REGION Network 181
   RUNG wire#powerrail
      Move(in := "Carrier_38_CarrierDriveAlarm", out1 => "DB_SDC_EMS_TA".EMS[38].TA[1].ALARM)
      wire#w1
      Move(in := "Carrier_38_CarrierDriveAlarm", out1 => "EMS".Carrier[38].SDC_IN.CarrierDriveAlarms)
   END_RUNG
   RUNG wire#powerrail
      Contact( "IndiconTempDebugON" )
   END_RUNG wire#w1
   // the same network as SCL:
   "DB_SDC_EMS_TA".EMS[38].TA[1].ALARM := "Carrier_38_CarrierDriveAlarm";
   IF TRUE OR "IndiconTempDebugON" THEN
       "EMS".Carrier[38].SDC_IN.CarrierDriveAlarms := "Carrier_38_CarrierDriveAlarm";
   END_IF;
END_REGION

REGION Network 182
   RUNG wire#powerrail
      Move(in := "Carrier_38_SDCFaultCode", out1 => "DB101_DB_SDC_FAULTS".Carrier_Fault[38])
      wire#w1
      Move(in := "Carrier_38_SDCFaultCode", out1 => "EMS".Carrier[38].SDC_IN.CarrierFaults)
   END_RUNG
   RUNG wire#powerrail
      Contact( "IndiconTempDebugON" )
   END_RUNG wire#w1
   // the same network as SCL:
   "DB101_DB_SDC_FAULTS".Carrier_Fault[38] := "Carrier_38_SDCFaultCode";
   IF TRUE OR "IndiconTempDebugON" THEN
       "EMS".Carrier[38].SDC_IN.CarrierFaults := "Carrier_38_SDCFaultCode";
   END_IF;
END_REGION

REGION Network 183
   RUNG wire#powerrail
      Contact( "Carrier_38_Status.5" )
      Coil( "EMS".Carrier[38].SDC_IN.RunningFWD )
   END_RUNG
   // the same network as SCL:
   "EMS".Carrier[38].SDC_IN.RunningFWD := "Carrier_38_Status.5";
END_REGION

REGION Network 184
   RUNG wire#powerrail
      Contact( "Carrier_38_Status.6" )
      Coil( "EMS".Carrier[38].SDC_IN.RunningREV )
   END_RUNG
   // the same network as SCL:
   "EMS".Carrier[38].SDC_IN.RunningREV := "Carrier_38_Status.6";
END_REGION

REGION Network 185
   RUNG wire#powerrail
      Contact( "Carrier_38_Status.7" )
      Coil( "EMS".Carrier[38].SDC_IN.IR_Remote_9_Pressed )
   END_RUNG
   // the same network as SCL:
   "EMS".Carrier[38].SDC_IN.IR_Remote_9_Pressed := "Carrier_38_Status.7";
END_REGION

REGION Network 186
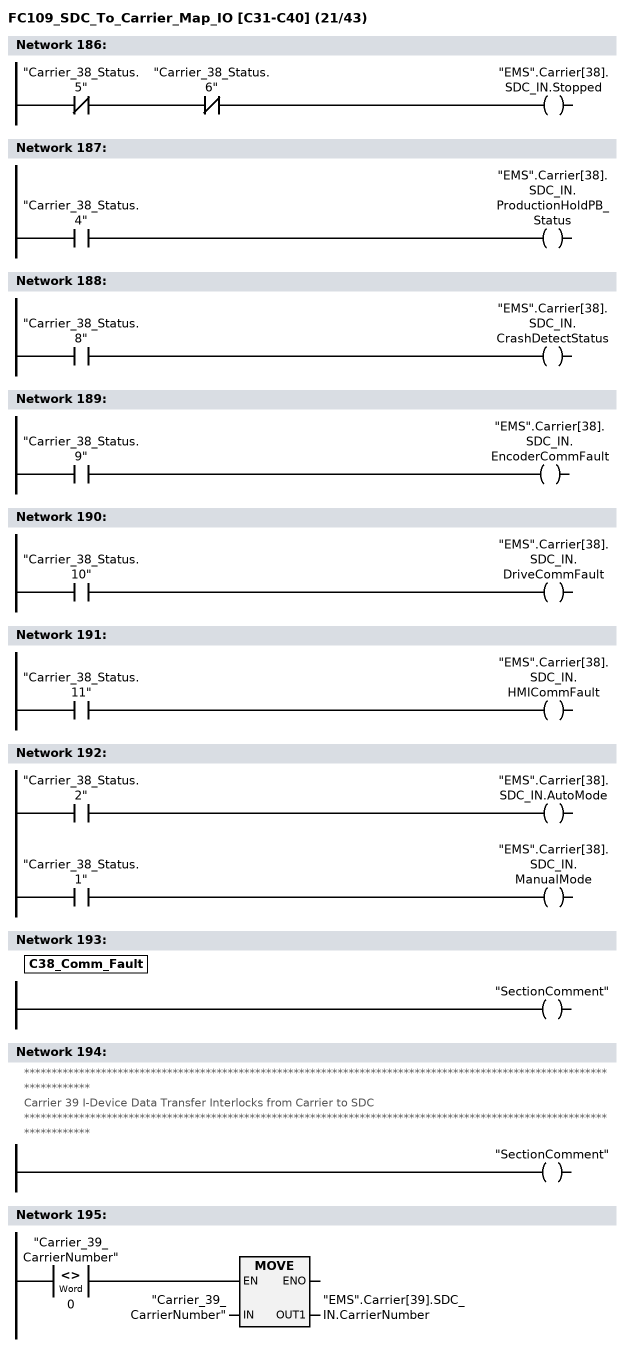
   RUNG wire#powerrail
      I_Contact( "Carrier_38_Status.5" )
      I_Contact( "Carrier_38_Status.6" )
      Coil( "EMS".Carrier[38].SDC_IN.Stopped )
   END_RUNG
   // the same network as SCL:
   "EMS".Carrier[38].SDC_IN.Stopped := NOT "Carrier_38_Status.5" AND NOT "Carrier_38_Status.6";
END_REGION

REGION Network 187
   RUNG wire#powerrail
      Contact( "Carrier_38_Status.4" )
      Coil( "EMS".Carrier[38].SDC_IN.ProductionHoldPB_Status )
   END_RUNG
   // the same network as SCL:
   "EMS".Carrier[38].SDC_IN.ProductionHoldPB_Status := "Carrier_38_Status.4";
END_REGION

REGION Network 188
   RUNG wire#powerrail
      Contact( "Carrier_38_Status.8" )
      Coil( "EMS".Carrier[38].SDC_IN.CrashDetectStatus )
   END_RUNG
   // the same network as SCL:
   "EMS".Carrier[38].SDC_IN.CrashDetectStatus := "Carrier_38_Status.8";
END_REGION

REGION Network 189
   RUNG wire#powerrail
      Contact( "Carrier_38_Status.9" )
      Coil( "EMS".Carrier[38].SDC_IN.EncoderCommFault )
   END_RUNG
   // the same network as SCL:
   "EMS".Carrier[38].SDC_IN.EncoderCommFault := "Carrier_38_Status.9";
END_REGION

REGION Network 190
   RUNG wire#powerrail
      Contact( "Carrier_38_Status.10" )
      Coil( "EMS".Carrier[38].SDC_IN.DriveCommFault )
   END_RUNG
   // the same network as SCL:
   "EMS".Carrier[38].SDC_IN.DriveCommFault := "Carrier_38_Status.10";
END_REGION

REGION Network 191
   RUNG wire#powerrail
      Contact( "Carrier_38_Status.11" )
      Coil( "EMS".Carrier[38].SDC_IN.HMICommFault )
   END_RUNG
   // the same network as SCL:
   "EMS".Carrier[38].SDC_IN.HMICommFault := "Carrier_38_Status.11";
END_REGION

REGION Network 192
   RUNG wire#powerrail
      Contact( "Carrier_38_Status.2" )
      Coil( "EMS".Carrier[38].SDC_IN.AutoMode )
   END_RUNG
   RUNG wire#powerrail
      Contact( "Carrier_38_Status.1" )
      Coil( "EMS".Carrier[38].SDC_IN.ManualMode )
   END_RUNG
   // the same network as SCL:
   "EMS".Carrier[38].SDC_IN.AutoMode := "Carrier_38_Status.2";
   "EMS".Carrier[38].SDC_IN.ManualMode := "Carrier_38_Status.1";
END_REGION

REGION Network 193
   Label( C38_Comm_Fault )
   RUNG wire#powerrail
      Coil( "SectionComment" )
   END_RUNG
   // the same network as SCL:
   C38_Comm_Fault:
   "SectionComment" := TRUE;
END_REGION

REGION Network 194
   // **********************************************************************************************************************
   // 
   // Carrier 39 I-Device Data Transfer Interlocks from Carrier to SDC
   // 
   // **********************************************************************************************************************
   RUNG wire#powerrail
      Coil( "SectionComment" )
   END_RUNG
   // the same network as SCL:
   "SectionComment" := TRUE;
END_REGION

REGION Network 195
   RUNG wire#powerrail
      { S7_Templates := "SrcType := Word" } NE_Contact(in1 := "Carrier_39_CarrierNumber", in2 := 0)
      Move(in := "Carrier_39_CarrierNumber", out1 => "EMS".Carrier[39].SDC_IN.CarrierNumber)
   END_RUNG
   // the same network as SCL:
   IF "Carrier_39_CarrierNumber" <> 0 THEN
       "EMS".Carrier[39].SDC_IN.CarrierNumber := "Carrier_39_CarrierNumber";
   END_IF;
END_REGION

REGION Network 196
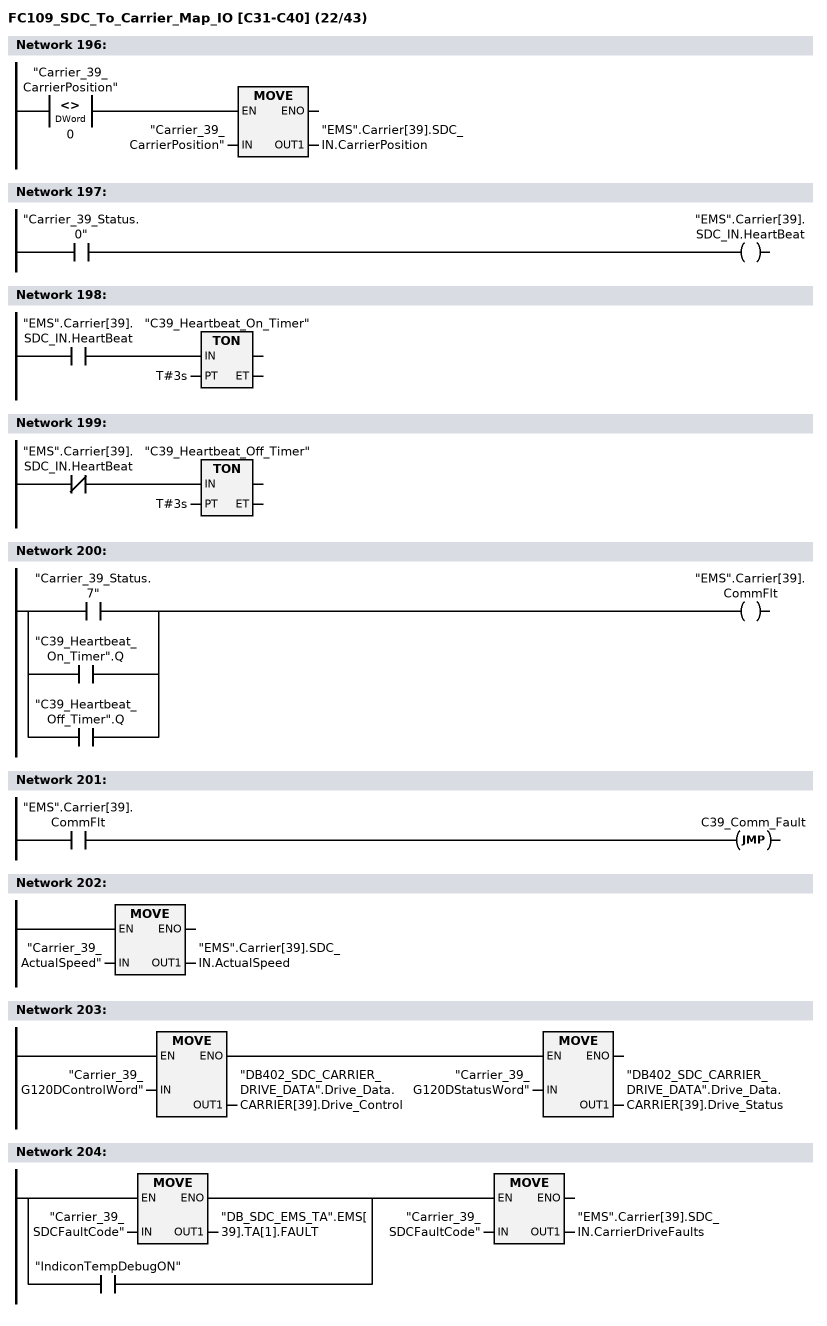
   RUNG wire#powerrail
      { S7_Templates := "SrcType := DWord" } NE_Contact(in1 := "Carrier_39_CarrierPosition", in2 := 0)
      Move(in := "Carrier_39_CarrierPosition", out1 => "EMS".Carrier[39].SDC_IN.CarrierPosition)
   END_RUNG
   // the same network as SCL:
   IF "Carrier_39_CarrierPosition" <> 0 THEN
       "EMS".Carrier[39].SDC_IN.CarrierPosition := "Carrier_39_CarrierPosition";
   END_IF;
END_REGION

REGION Network 197
   RUNG wire#powerrail
      Contact( "Carrier_39_Status.0" )
      Coil( "EMS".Carrier[39].SDC_IN.HeartBeat )
   END_RUNG
   // the same network as SCL:
   "EMS".Carrier[39].SDC_IN.HeartBeat := "Carrier_39_Status.0";
END_REGION

REGION Network 198
   "C39_Heartbeat_On_Timer".TON(IN := "EMS".Carrier[39].SDC_IN.HeartBeat, PT := T#3s);
END_REGION

REGION Network 199
   "C39_Heartbeat_Off_Timer".TON(IN := NOT "EMS".Carrier[39].SDC_IN.HeartBeat, PT := T#3s);
END_REGION

REGION Network 200
   RUNG wire#powerrail
      Contact( "Carrier_39_Status.7" )
      wire#w1
      Coil( "EMS".Carrier[39].CommFlt )
   END_RUNG
   RUNG wire#powerrail
      Contact( "C39_Heartbeat_On_Timer".Q )
   END_RUNG wire#w1
   RUNG wire#powerrail
      Contact( "C39_Heartbeat_Off_Timer".Q )
   END_RUNG wire#w1
   // the same network as SCL:
   "EMS".Carrier[39].CommFlt := "Carrier_39_Status.7" OR "C39_Heartbeat_On_Timer".Q OR "C39_Heartbeat_Off_Timer".Q;
END_REGION

REGION Network 201
   RUNG wire#powerrail
      Contact( "EMS".Carrier[39].CommFlt )
      JumpCoil( C39_Comm_Fault )
   END_RUNG
   // the same network as SCL:
   IF "EMS".Carrier[39].CommFlt THEN GOTO C39_Comm_Fault; END_IF;
END_REGION

REGION Network 202
   RUNG wire#powerrail
      Move(in := "Carrier_39_ActualSpeed", out1 => "EMS".Carrier[39].SDC_IN.ActualSpeed)
   END_RUNG
   // the same network as SCL:
   "EMS".Carrier[39].SDC_IN.ActualSpeed := "Carrier_39_ActualSpeed";
END_REGION

REGION Network 203
   RUNG wire#powerrail
      Move(in := "Carrier_39_G120DControlWord", out1 => "DB402_SDC_CARRIER_DRIVE_DATA".Drive_Data.CARRIER[39].Drive_Control)
      Move(in := "Carrier_39_G120DStatusWord", out1 => "DB402_SDC_CARRIER_DRIVE_DATA".Drive_Data.CARRIER[39].Drive_Status)
   END_RUNG
   // the same network as SCL:
   "DB402_SDC_CARRIER_DRIVE_DATA".Drive_Data.CARRIER[39].Drive_Control := "Carrier_39_G120DControlWord";
   "DB402_SDC_CARRIER_DRIVE_DATA".Drive_Data.CARRIER[39].Drive_Status := "Carrier_39_G120DStatusWord";
END_REGION

REGION Network 204
   RUNG wire#powerrail
      Move(in := "Carrier_39_SDCFaultCode", out1 => "DB_SDC_EMS_TA".EMS[39].TA[1].FAULT)
      wire#w1
      Move(in := "Carrier_39_SDCFaultCode", out1 => "EMS".Carrier[39].SDC_IN.CarrierDriveFaults)
   END_RUNG
   RUNG wire#powerrail
      Contact( "IndiconTempDebugON" )
   END_RUNG wire#w1
   // the same network as SCL:
   "DB_SDC_EMS_TA".EMS[39].TA[1].FAULT := "Carrier_39_SDCFaultCode";
   IF TRUE OR "IndiconTempDebugON" THEN
       "EMS".Carrier[39].SDC_IN.CarrierDriveFaults := "Carrier_39_SDCFaultCode";
   END_IF;
END_REGION

REGION Network 205
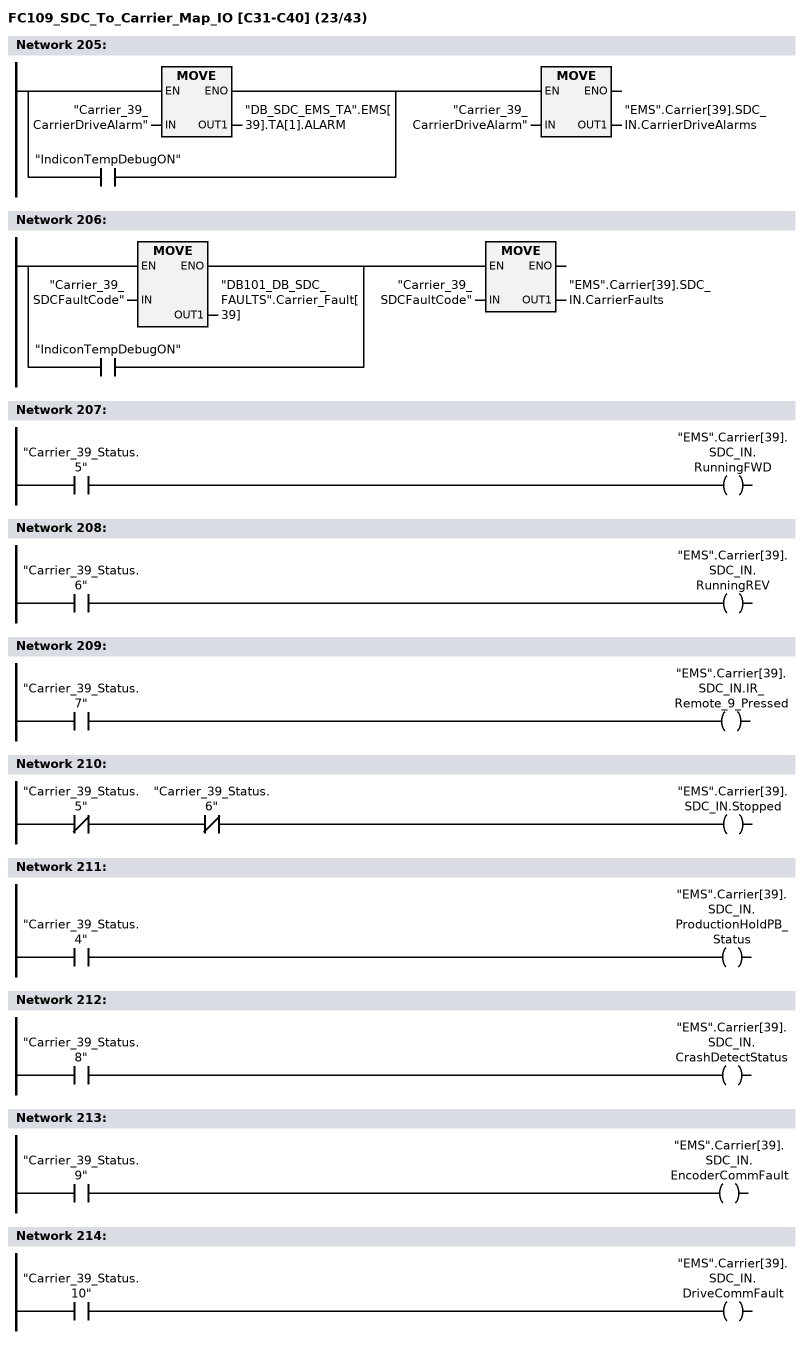
   RUNG wire#powerrail
      Move(in := "Carrier_39_CarrierDriveAlarm", out1 => "DB_SDC_EMS_TA".EMS[39].TA[1].ALARM)
      wire#w1
      Move(in := "Carrier_39_CarrierDriveAlarm", out1 => "EMS".Carrier[39].SDC_IN.CarrierDriveAlarms)
   END_RUNG
   RUNG wire#powerrail
      Contact( "IndiconTempDebugON" )
   END_RUNG wire#w1
   // the same network as SCL:
   "DB_SDC_EMS_TA".EMS[39].TA[1].ALARM := "Carrier_39_CarrierDriveAlarm";
   IF TRUE OR "IndiconTempDebugON" THEN
       "EMS".Carrier[39].SDC_IN.CarrierDriveAlarms := "Carrier_39_CarrierDriveAlarm";
   END_IF;
END_REGION

REGION Network 206
   RUNG wire#powerrail
      Move(in := "Carrier_39_SDCFaultCode", out1 => "DB101_DB_SDC_FAULTS".Carrier_Fault[39])
      wire#w1
      Move(in := "Carrier_39_SDCFaultCode", out1 => "EMS".Carrier[39].SDC_IN.CarrierFaults)
   END_RUNG
   RUNG wire#powerrail
      Contact( "IndiconTempDebugON" )
   END_RUNG wire#w1
   // the same network as SCL:
   "DB101_DB_SDC_FAULTS".Carrier_Fault[39] := "Carrier_39_SDCFaultCode";
   IF TRUE OR "IndiconTempDebugON" THEN
       "EMS".Carrier[39].SDC_IN.CarrierFaults := "Carrier_39_SDCFaultCode";
   END_IF;
END_REGION

REGION Network 207
   RUNG wire#powerrail
      Contact( "Carrier_39_Status.5" )
      Coil( "EMS".Carrier[39].SDC_IN.RunningFWD )
   END_RUNG
   // the same network as SCL:
   "EMS".Carrier[39].SDC_IN.RunningFWD := "Carrier_39_Status.5";
END_REGION

REGION Network 208
   RUNG wire#powerrail
      Contact( "Carrier_39_Status.6" )
      Coil( "EMS".Carrier[39].SDC_IN.RunningREV )
   END_RUNG
   // the same network as SCL:
   "EMS".Carrier[39].SDC_IN.RunningREV := "Carrier_39_Status.6";
END_REGION

REGION Network 209
   RUNG wire#powerrail
      Contact( "Carrier_39_Status.7" )
      Coil( "EMS".Carrier[39].SDC_IN.IR_Remote_9_Pressed )
   END_RUNG
   // the same network as SCL:
   "EMS".Carrier[39].SDC_IN.IR_Remote_9_Pressed := "Carrier_39_Status.7";
END_REGION

REGION Network 210
   RUNG wire#powerrail
      I_Contact( "Carrier_39_Status.5" )
      I_Contact( "Carrier_39_Status.6" )
      Coil( "EMS".Carrier[39].SDC_IN.Stopped )
   END_RUNG
   // the same network as SCL:
   "EMS".Carrier[39].SDC_IN.Stopped := NOT "Carrier_39_Status.5" AND NOT "Carrier_39_Status.6";
END_REGION

REGION Network 211
   RUNG wire#powerrail
      Contact( "Carrier_39_Status.4" )
      Coil( "EMS".Carrier[39].SDC_IN.ProductionHoldPB_Status )
   END_RUNG
   // the same network as SCL:
   "EMS".Carrier[39].SDC_IN.ProductionHoldPB_Status := "Carrier_39_Status.4";
END_REGION

REGION Network 212
   RUNG wire#powerrail
      Contact( "Carrier_39_Status.8" )
      Coil( "EMS".Carrier[39].SDC_IN.CrashDetectStatus )
   END_RUNG
   // the same network as SCL:
   "EMS".Carrier[39].SDC_IN.CrashDetectStatus := "Carrier_39_Status.8";
END_REGION

REGION Network 213
   RUNG wire#powerrail
      Contact( "Carrier_39_Status.9" )
      Coil( "EMS".Carrier[39].SDC_IN.EncoderCommFault )
   END_RUNG
   // the same network as SCL:
   "EMS".Carrier[39].SDC_IN.EncoderCommFault := "Carrier_39_Status.9";
END_REGION

REGION Network 214
   RUNG wire#powerrail
      Contact( "Carrier_39_Status.10" )
      Coil( "EMS".Carrier[39].SDC_IN.DriveCommFault )
   END_RUNG
   // the same network as SCL:
   "EMS".Carrier[39].SDC_IN.DriveCommFault := "Carrier_39_Status.10";
END_REGION

REGION Network 215
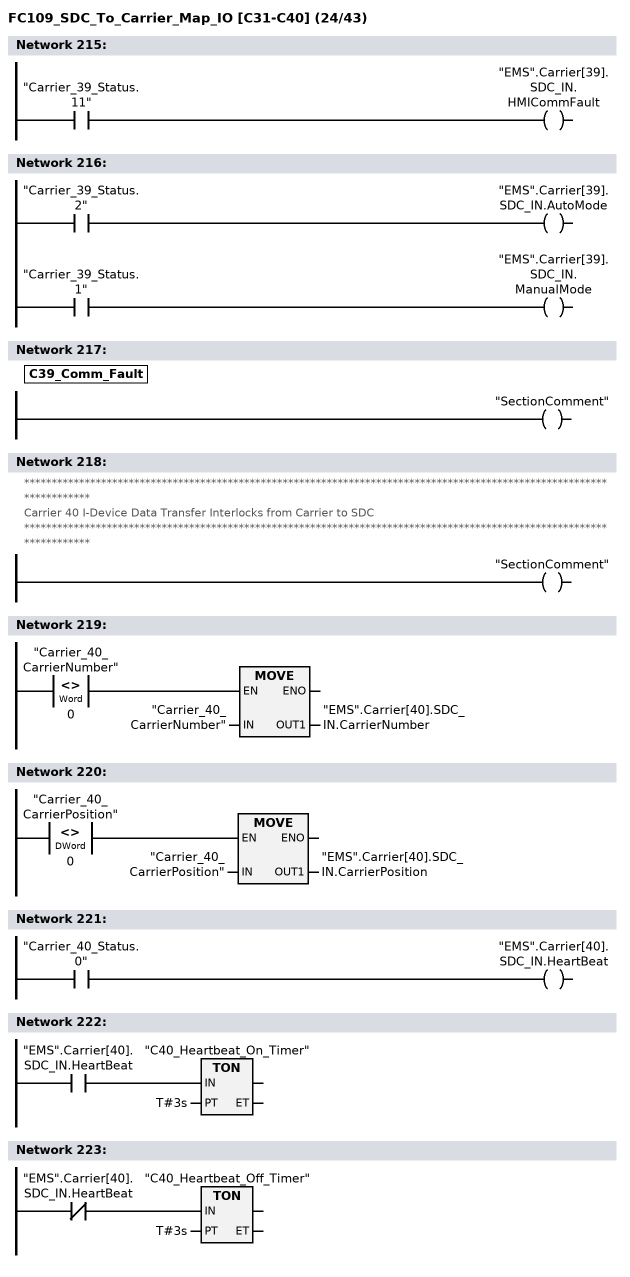
   RUNG wire#powerrail
      Contact( "Carrier_39_Status.11" )
      Coil( "EMS".Carrier[39].SDC_IN.HMICommFault )
   END_RUNG
   // the same network as SCL:
   "EMS".Carrier[39].SDC_IN.HMICommFault := "Carrier_39_Status.11";
END_REGION

REGION Network 216
   RUNG wire#powerrail
      Contact( "Carrier_39_Status.2" )
      Coil( "EMS".Carrier[39].SDC_IN.AutoMode )
   END_RUNG
   RUNG wire#powerrail
      Contact( "Carrier_39_Status.1" )
      Coil( "EMS".Carrier[39].SDC_IN.ManualMode )
   END_RUNG
   // the same network as SCL:
   "EMS".Carrier[39].SDC_IN.AutoMode := "Carrier_39_Status.2";
   "EMS".Carrier[39].SDC_IN.ManualMode := "Carrier_39_Status.1";
END_REGION

REGION Network 217
   Label( C39_Comm_Fault )
   RUNG wire#powerrail
      Coil( "SectionComment" )
   END_RUNG
   // the same network as SCL:
   C39_Comm_Fault:
   "SectionComment" := TRUE;
END_REGION

REGION Network 218
   // **********************************************************************************************************************
   // 
   // Carrier 40 I-Device Data Transfer Interlocks from Carrier to SDC
   // 
   // **********************************************************************************************************************
   RUNG wire#powerrail
      Coil( "SectionComment" )
   END_RUNG
   // the same network as SCL:
   "SectionComment" := TRUE;
END_REGION

REGION Network 219
   RUNG wire#powerrail
      { S7_Templates := "SrcType := Word" } NE_Contact(in1 := "Carrier_40_CarrierNumber", in2 := 0)
      Move(in := "Carrier_40_CarrierNumber", out1 => "EMS".Carrier[40].SDC_IN.CarrierNumber)
   END_RUNG
   // the same network as SCL:
   IF "Carrier_40_CarrierNumber" <> 0 THEN
       "EMS".Carrier[40].SDC_IN.CarrierNumber := "Carrier_40_CarrierNumber";
   END_IF;
END_REGION

REGION Network 220
   RUNG wire#powerrail
      { S7_Templates := "SrcType := DWord" } NE_Contact(in1 := "Carrier_40_CarrierPosition", in2 := 0)
      Move(in := "Carrier_40_CarrierPosition", out1 => "EMS".Carrier[40].SDC_IN.CarrierPosition)
   END_RUNG
   // the same network as SCL:
   IF "Carrier_40_CarrierPosition" <> 0 THEN
       "EMS".Carrier[40].SDC_IN.CarrierPosition := "Carrier_40_CarrierPosition";
   END_IF;
END_REGION

REGION Network 221
   RUNG wire#powerrail
      Contact( "Carrier_40_Status.0" )
      Coil( "EMS".Carrier[40].SDC_IN.HeartBeat )
   END_RUNG
   // the same network as SCL:
   "EMS".Carrier[40].SDC_IN.HeartBeat := "Carrier_40_Status.0";
END_REGION

REGION Network 222
   "C40_Heartbeat_On_Timer".TON(IN := "EMS".Carrier[40].SDC_IN.HeartBeat, PT := T#3s);
END_REGION

REGION Network 223
   "C40_Heartbeat_Off_Timer".TON(IN := NOT "EMS".Carrier[40].SDC_IN.HeartBeat, PT := T#3s);
END_REGION

REGION Network 224
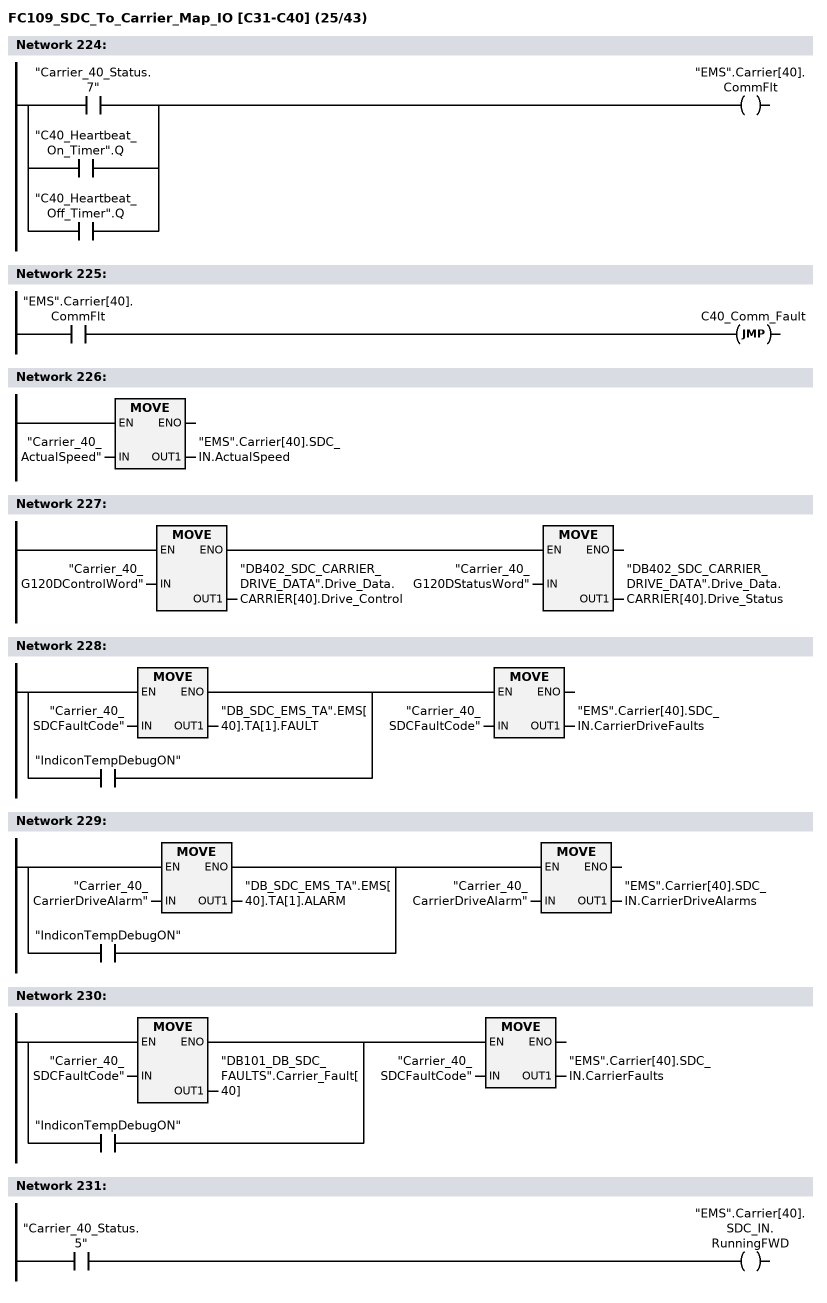
   RUNG wire#powerrail
      Contact( "Carrier_40_Status.7" )
      wire#w1
      Coil( "EMS".Carrier[40].CommFlt )
   END_RUNG
   RUNG wire#powerrail
      Contact( "C40_Heartbeat_On_Timer".Q )
   END_RUNG wire#w1
   RUNG wire#powerrail
      Contact( "C40_Heartbeat_Off_Timer".Q )
   END_RUNG wire#w1
   // the same network as SCL:
   "EMS".Carrier[40].CommFlt := "Carrier_40_Status.7" OR "C40_Heartbeat_On_Timer".Q OR "C40_Heartbeat_Off_Timer".Q;
END_REGION

REGION Network 225
   RUNG wire#powerrail
      Contact( "EMS".Carrier[40].CommFlt )
      JumpCoil( C40_Comm_Fault )
   END_RUNG
   // the same network as SCL:
   IF "EMS".Carrier[40].CommFlt THEN GOTO C40_Comm_Fault; END_IF;
END_REGION

REGION Network 226
   RUNG wire#powerrail
      Move(in := "Carrier_40_ActualSpeed", out1 => "EMS".Carrier[40].SDC_IN.ActualSpeed)
   END_RUNG
   // the same network as SCL:
   "EMS".Carrier[40].SDC_IN.ActualSpeed := "Carrier_40_ActualSpeed";
END_REGION

REGION Network 227
   RUNG wire#powerrail
      Move(in := "Carrier_40_G120DControlWord", out1 => "DB402_SDC_CARRIER_DRIVE_DATA".Drive_Data.CARRIER[40].Drive_Control)
      Move(in := "Carrier_40_G120DStatusWord", out1 => "DB402_SDC_CARRIER_DRIVE_DATA".Drive_Data.CARRIER[40].Drive_Status)
   END_RUNG
   // the same network as SCL:
   "DB402_SDC_CARRIER_DRIVE_DATA".Drive_Data.CARRIER[40].Drive_Control := "Carrier_40_G120DControlWord";
   "DB402_SDC_CARRIER_DRIVE_DATA".Drive_Data.CARRIER[40].Drive_Status := "Carrier_40_G120DStatusWord";
END_REGION

REGION Network 228
   RUNG wire#powerrail
      Move(in := "Carrier_40_SDCFaultCode", out1 => "DB_SDC_EMS_TA".EMS[40].TA[1].FAULT)
      wire#w1
      Move(in := "Carrier_40_SDCFaultCode", out1 => "EMS".Carrier[40].SDC_IN.CarrierDriveFaults)
   END_RUNG
   RUNG wire#powerrail
      Contact( "IndiconTempDebugON" )
   END_RUNG wire#w1
   // the same network as SCL:
   "DB_SDC_EMS_TA".EMS[40].TA[1].FAULT := "Carrier_40_SDCFaultCode";
   IF TRUE OR "IndiconTempDebugON" THEN
       "EMS".Carrier[40].SDC_IN.CarrierDriveFaults := "Carrier_40_SDCFaultCode";
   END_IF;
END_REGION

REGION Network 229
   RUNG wire#powerrail
      Move(in := "Carrier_40_CarrierDriveAlarm", out1 => "DB_SDC_EMS_TA".EMS[40].TA[1].ALARM)
      wire#w1
      Move(in := "Carrier_40_CarrierDriveAlarm", out1 => "EMS".Carrier[40].SDC_IN.CarrierDriveAlarms)
   END_RUNG
   RUNG wire#powerrail
      Contact( "IndiconTempDebugON" )
   END_RUNG wire#w1
   // the same network as SCL:
   "DB_SDC_EMS_TA".EMS[40].TA[1].ALARM := "Carrier_40_CarrierDriveAlarm";
   IF TRUE OR "IndiconTempDebugON" THEN
       "EMS".Carrier[40].SDC_IN.CarrierDriveAlarms := "Carrier_40_CarrierDriveAlarm";
   END_IF;
END_REGION

REGION Network 230
   RUNG wire#powerrail
      Move(in := "Carrier_40_SDCFaultCode", out1 => "DB101_DB_SDC_FAULTS".Carrier_Fault[40])
      wire#w1
      Move(in := "Carrier_40_SDCFaultCode", out1 => "EMS".Carrier[40].SDC_IN.CarrierFaults)
   END_RUNG
   RUNG wire#powerrail
      Contact( "IndiconTempDebugON" )
   END_RUNG wire#w1
   // the same network as SCL:
   "DB101_DB_SDC_FAULTS".Carrier_Fault[40] := "Carrier_40_SDCFaultCode";
   IF TRUE OR "IndiconTempDebugON" THEN
       "EMS".Carrier[40].SDC_IN.CarrierFaults := "Carrier_40_SDCFaultCode";
   END_IF;
END_REGION

REGION Network 231
   RUNG wire#powerrail
      Contact( "Carrier_40_Status.5" )
      Coil( "EMS".Carrier[40].SDC_IN.RunningFWD )
   END_RUNG
   // the same network as SCL:
   "EMS".Carrier[40].SDC_IN.RunningFWD := "Carrier_40_Status.5";
END_REGION

REGION Network 232
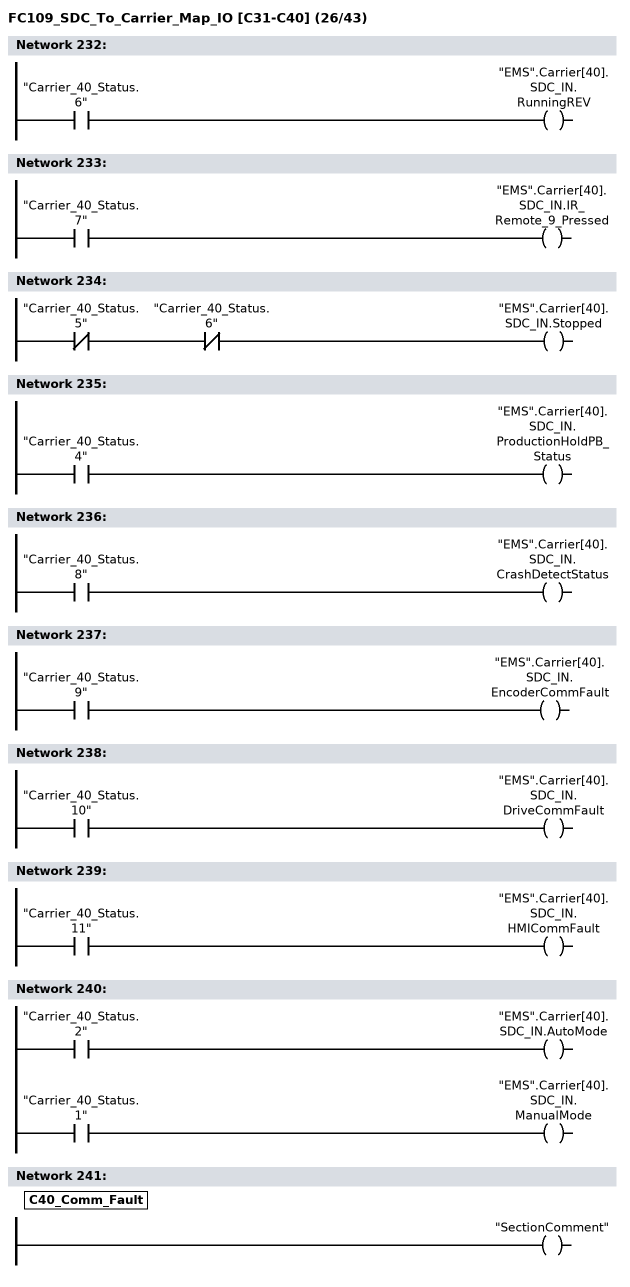
   RUNG wire#powerrail
      Contact( "Carrier_40_Status.6" )
      Coil( "EMS".Carrier[40].SDC_IN.RunningREV )
   END_RUNG
   // the same network as SCL:
   "EMS".Carrier[40].SDC_IN.RunningREV := "Carrier_40_Status.6";
END_REGION

REGION Network 233
   RUNG wire#powerrail
      Contact( "Carrier_40_Status.7" )
      Coil( "EMS".Carrier[40].SDC_IN.IR_Remote_9_Pressed )
   END_RUNG
   // the same network as SCL:
   "EMS".Carrier[40].SDC_IN.IR_Remote_9_Pressed := "Carrier_40_Status.7";
END_REGION

REGION Network 234
   RUNG wire#powerrail
      I_Contact( "Carrier_40_Status.5" )
      I_Contact( "Carrier_40_Status.6" )
      Coil( "EMS".Carrier[40].SDC_IN.Stopped )
   END_RUNG
   // the same network as SCL:
   "EMS".Carrier[40].SDC_IN.Stopped := NOT "Carrier_40_Status.5" AND NOT "Carrier_40_Status.6";
END_REGION

REGION Network 235
   RUNG wire#powerrail
      Contact( "Carrier_40_Status.4" )
      Coil( "EMS".Carrier[40].SDC_IN.ProductionHoldPB_Status )
   END_RUNG
   // the same network as SCL:
   "EMS".Carrier[40].SDC_IN.ProductionHoldPB_Status := "Carrier_40_Status.4";
END_REGION

REGION Network 236
   RUNG wire#powerrail
      Contact( "Carrier_40_Status.8" )
      Coil( "EMS".Carrier[40].SDC_IN.CrashDetectStatus )
   END_RUNG
   // the same network as SCL:
   "EMS".Carrier[40].SDC_IN.CrashDetectStatus := "Carrier_40_Status.8";
END_REGION

REGION Network 237
   RUNG wire#powerrail
      Contact( "Carrier_40_Status.9" )
      Coil( "EMS".Carrier[40].SDC_IN.EncoderCommFault )
   END_RUNG
   // the same network as SCL:
   "EMS".Carrier[40].SDC_IN.EncoderCommFault := "Carrier_40_Status.9";
END_REGION

REGION Network 238
   RUNG wire#powerrail
      Contact( "Carrier_40_Status.10" )
      Coil( "EMS".Carrier[40].SDC_IN.DriveCommFault )
   END_RUNG
   // the same network as SCL:
   "EMS".Carrier[40].SDC_IN.DriveCommFault := "Carrier_40_Status.10";
END_REGION

REGION Network 239
   RUNG wire#powerrail
      Contact( "Carrier_40_Status.11" )
      Coil( "EMS".Carrier[40].SDC_IN.HMICommFault )
   END_RUNG
   // the same network as SCL:
   "EMS".Carrier[40].SDC_IN.HMICommFault := "Carrier_40_Status.11";
END_REGION

REGION Network 240
   RUNG wire#powerrail
      Contact( "Carrier_40_Status.2" )
      Coil( "EMS".Carrier[40].SDC_IN.AutoMode )
   END_RUNG
   RUNG wire#powerrail
      Contact( "Carrier_40_Status.1" )
      Coil( "EMS".Carrier[40].SDC_IN.ManualMode )
   END_RUNG
   // the same network as SCL:
   "EMS".Carrier[40].SDC_IN.AutoMode := "Carrier_40_Status.2";
   "EMS".Carrier[40].SDC_IN.ManualMode := "Carrier_40_Status.1";
END_REGION

REGION Network 241
   Label( C40_Comm_Fault )
   RUNG wire#powerrail
      Coil( "SectionComment" )
   END_RUNG
   // the same network as SCL:
   C40_Comm_Fault:
   "SectionComment" := TRUE;
END_REGION

REGION Network 242
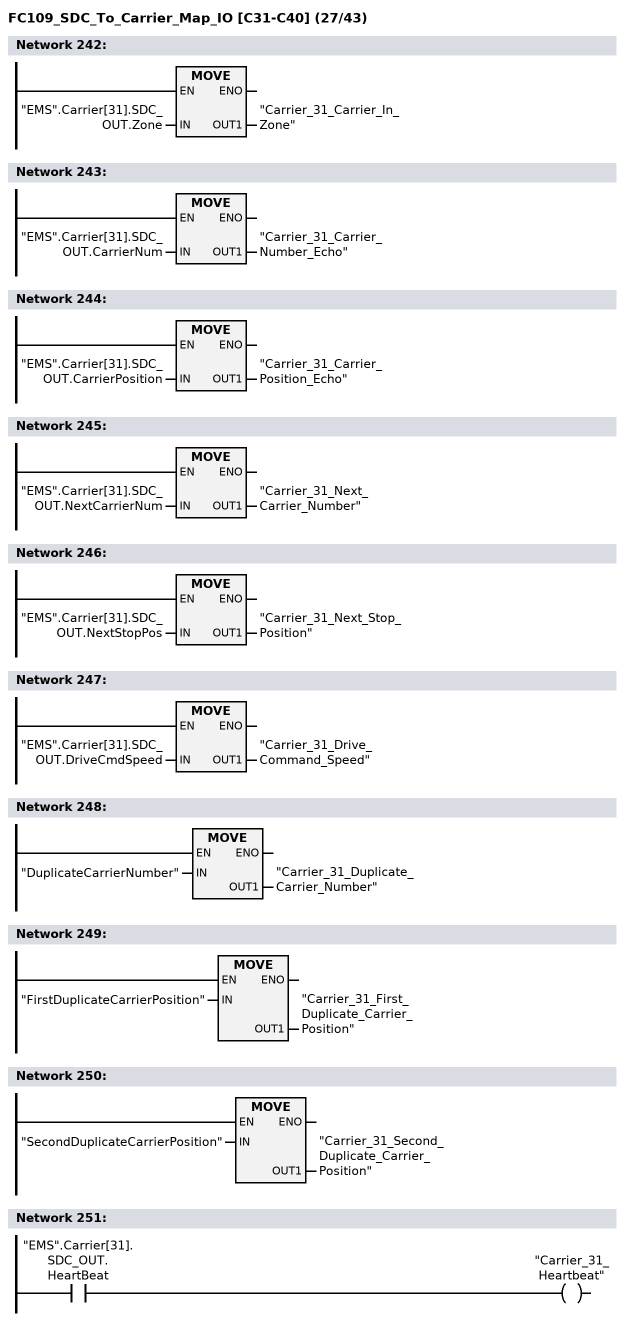
   RUNG wire#powerrail
      Move(in := "EMS".Carrier[31].SDC_OUT.Zone, out1 => "Carrier_31_Carrier_In_Zone")
   END_RUNG
   // the same network as SCL:
   "Carrier_31_Carrier_In_Zone" := "EMS".Carrier[31].SDC_OUT.Zone;
END_REGION

REGION Network 243
   RUNG wire#powerrail
      Move(in := "EMS".Carrier[31].SDC_OUT.CarrierNum, out1 => "Carrier_31_Carrier_Number_Echo")
   END_RUNG
   // the same network as SCL:
   "Carrier_31_Carrier_Number_Echo" := "EMS".Carrier[31].SDC_OUT.CarrierNum;
END_REGION

REGION Network 244
   RUNG wire#powerrail
      Move(in := "EMS".Carrier[31].SDC_OUT.CarrierPosition, out1 => "Carrier_31_Carrier_Position_Echo")
   END_RUNG
   // the same network as SCL:
   "Carrier_31_Carrier_Position_Echo" := "EMS".Carrier[31].SDC_OUT.CarrierPosition;
END_REGION

REGION Network 245
   RUNG wire#powerrail
      Move(in := "EMS".Carrier[31].SDC_OUT.NextCarrierNum, out1 => "Carrier_31_Next_Carrier_Number")
   END_RUNG
   // the same network as SCL:
   "Carrier_31_Next_Carrier_Number" := "EMS".Carrier[31].SDC_OUT.NextCarrierNum;
END_REGION

REGION Network 246
   RUNG wire#powerrail
      Move(in := "EMS".Carrier[31].SDC_OUT.NextStopPos, out1 => "Carrier_31_Next_Stop_Position")
   END_RUNG
   // the same network as SCL:
   "Carrier_31_Next_Stop_Position" := "EMS".Carrier[31].SDC_OUT.NextStopPos;
END_REGION

REGION Network 247
   RUNG wire#powerrail
      Move(in := "EMS".Carrier[31].SDC_OUT.DriveCmdSpeed, out1 => "Carrier_31_Drive_Command_Speed")
   END_RUNG
   // the same network as SCL:
   "Carrier_31_Drive_Command_Speed" := "EMS".Carrier[31].SDC_OUT.DriveCmdSpeed;
END_REGION

REGION Network 248
   RUNG wire#powerrail
      Move(in := "DuplicateCarrierNumber", out1 => "Carrier_31_Duplicate_Carrier_Number")
   END_RUNG
   // the same network as SCL:
   "Carrier_31_Duplicate_Carrier_Number" := "DuplicateCarrierNumber";
END_REGION

REGION Network 249
   RUNG wire#powerrail
      Move(in := "FirstDuplicateCarrierPosition", out1 => "Carrier_31_First_Duplicate_Carrier_Position")
   END_RUNG
   // the same network as SCL:
   "Carrier_31_First_Duplicate_Carrier_Position" := "FirstDuplicateCarrierPosition";
END_REGION

REGION Network 250
   RUNG wire#powerrail
      Move(in := "SecondDuplicateCarrierPosition", out1 => "Carrier_31_Second_Duplicate_Carrier_Position")
   END_RUNG
   // the same network as SCL:
   "Carrier_31_Second_Duplicate_Carrier_Position" := "SecondDuplicateCarrierPosition";
END_REGION

REGION Network 251
   RUNG wire#powerrail
      Contact( "EMS".Carrier[31].SDC_OUT.HeartBeat )
      Coil( "Carrier_31_Heartbeat" )
   END_RUNG
   // the same network as SCL:
   "Carrier_31_Heartbeat" := "EMS".Carrier[31].SDC_OUT.HeartBeat;
END_REGION

REGION Network 252